(* Logix 5000 project; controller Joltek_RA_5069PLC002 vendor 1 type 14 code 226 rev 34.15; software revision 34.04 *)

TASK MainTask (continuous, watchdog 500 ms) : MainProgram
TASK SafetyTask (periodic, rate 20 ms, priority 10, watchdog 20 ms, safety) : SafetyProgram

MODULES
   Local : vendor 1 type 14 code 226 (5069 0, rev 34.15)
      Joltek_SW001 : vendor 1 type 12 code 231 (Ethernet 192.168.1.70, rev 13.8, Output RPI 1000 ms)
END_MODULES

TYPE UDT_ErrorDataLog :
STRUCT
   Time : UDT_Timestamp;
   DINTlog : DINT[10];
   REALlog : REAL[10];
END_STRUCT
END_TYPE

TYPE UDT_Line :
STRUCT
   Filler : UDT_Machine;
   Capper : UDT_Machine;
   Labeler : UDT_Machine;
   CasePAcker : UDT_Machine;
END_STRUCT
END_TYPE

TYPE UDT_Machine :
STRUCT
   Status : INT;
   Running : TIMER;
   Running_B : BOOL;
   CustomData : DINT[10];
   CustomREALData : REAL[10];
   Faulted : DINT;
END_STRUCT
END_TYPE

TYPE UDT_Timestamp :
STRUCT
   Year : DINT;
   Month : DINT;
   Day : DINT;
   Hour : DINT;
   Minute : DINT;
   Second : DINT;
END_STRUCT
END_TYPE

VAR_GLOBAL   (* controller tags *)
   FillerData : UDT_Machine;
   HMI_BOOL1 : BOOL[128] := ([0] := 1);
        [2]   // Filler - HMI | Station 1 Filling
        [3]   // Filler - HMI | Station 2 Filling
   HMI_INT : INT[100] := ([0] := 3, [1] := 717, [2] := 50, [3] := 16656, [5] := 10, [10] := 3, [11] := 85, [12] := 164, [14] := 9, [20] := 4, [21] := 115, [22] := 5, [23] := 9, [30] := 2, [31] := 66, [33] := 4100, [40] := 2, [41] := 8, [42] := 38, [50] := 4);
        [3].12   // Filler - Start Permissive
        [3].13   // Filler HMI - Start Command
        [23].0   // Labeler - Labeling in Process
        [23].1   // Labeler - Start Permissive
        [23].2   // Labeler - HMI Start Command
        [23].3   // Labeler - Stop Permissive
        [23].4   // Labeler - HMI Stop Command
        [23].5   // Labeler - HMI Faulted Status
        [23].6   // Labeler - HMI Fault Reset Command
        [33].0   // Case Packer - HMI | Case Folding in Progress
        [33].1   // Case Packer - HMI | Case Gluing in Progress
        [33].10   // Case Packer - HMI | Start Permissive
        [33].11   // Case Packer - HMI | Start Command
        [33].12   // Case Packer - HMI | Stop Permissive
        [33].13   // Case Packer - HMI | Stop Command
        [33].15   // Case Packer - HMI | Clear Fault Command
        [41].0   // Palletizer - HMI | Currently Palletizing
        [41].1   // Palletizer - HMI | Start Permissive
        [41].2   // Palletizer - HMI | Start Command
        [41].7   // Palletizer - HMI | Clear Pallet Command
        [50].0   // Line - HIM | Start Permissive
        [50].1   // Line - HIM | Start Command
        [50].2   // Line - HIM | Stop Permissive
        [50].3   // Line - HIM | Stop Command
        [50].5   // Line - HIM | Fault Reset Command
        [14].2   // Capper - HMI | Start Command
        [14].4   // Capper - HMI | Stop Command
        [14].6   // Capper - HMI | Fault Reset Command
   HMI_REAL : REAL[100] := ([0] := 100.0, [1] := 100.0, [2] := 100.0, [3] := 60.0, [4] := 42.0);
   Line1 : UDT_Line;
   Line34Pump3Motor342DischargeOfTank23_Sig : DINT;
   Line45Pump3MTR345InfeedRawIngredientFlou : DINT;
   Line6Pump1DischargeOfTank3 : DINT;
   Sys_DINT : DINT[100] := ([0] := 3, [1] := 3387, [2] := 6708, [3] := 68, [4] := 717, [5] := 10000, [6] := 10000, [7] := 1, [8] := 1, [9] := 1, [10] := 1, [11] := 1, [12] := 1, [13] := 1, [14] := 1, [15] := 1, [16] := 1, [17] := 1, [18] := 1, [19] := 1, [20] := 1, [21] := 1, [22] := 1, [23] := 1, [24] := 1, [25] := 1, [26] := 1, [27] := 1, [28] := 1, [29] := 1, [30] := 1, [31] := 1, [32] := 1, [33] := 1, [34] := 1, [35] := 1, [36] := 1, [39] := 50, [40] := 52, [41] := 10000, [42] := 85, [43] := 164, [44] := 20, [45] := 6100, [46] := 5, [47] := 115, [48] := 4, [49] := 66, [51] := 4200, [54] := 1, [55] := 4, [57] := 38);
        [0]   // Line 1 Motor 324 of the Conveyor 23 Discharge Pump 4-20mA Signal
        [1]   // Line 2 Motor 32334 of the Conveyor 2233 Discharge Pump 0-20mA Signal SCALED
        [3].1   // Filler - Stop
        [3].3   // Filler - Faulted
        [3].2   // Filler - Running
        [40].4   // Capper - Start Capping Process
        [4]   // Filler - Infeed Empty Bottle Count
        [3].0   // Filler - Start
        [3].4   // Filler - Alarm | Infeed Empty Bottle Conveyor Empty
        [3].5   // Filler - Alarm | Infeed Empty Bottle Conveyor Low
        [3].6   // Filler - Alarm | Discharge Filled Bottle Conveyor Full
        [3].7   // Filler - Alarm | Discharge Filled Bottle Conveyor Almost Full
        [40].2   // Capper - Running
        [40].5   // Capper Discharge Conveyor Full
        [40].6   // Capper Discharge Conveyor Almost Full
        [40].7   // Capper Infeed Conveyor Empty
        [40].8   // Capper Infeed Conveyor Almost Empty
        [44].0   // Labeler - Start
        [44].2   // Labeler - Running
        [39]   // Filled Bottle Conveyor Count
        [44].1   // Labeler - Stop
        [44].3   // Labeler - Faulted
        [43]   // Capper - Caps available in the hopper
        [44].5   // Labeler - Labeled Bottle Conveyor Full
        [44].6   // Labeler - Labeled Bottle Conveyor Almost Full
        [44].7   // Labeler - Capped Bottle Conveyor Empty
        [44].8   // Labeler - Capped Bottle Conveyor Almost Empty
        [44].9   // Labeler - Unwind Station Empty
        [44].10   // Labeler - Unwind Station Almost Empty
        [48].0   // Case Packer - Start
        [48].1   // Case Packer - Stop
        [48].3   // Case Packer - Faulted
        [48].2   // Case Packer - Running
        [48].4   // Case Packer - Case Filling Station
        [46]   // Labeled Bollte Conveyor Count
        [49]   // Case Packer - Empty Case Count
        [48].5   // Case Packer - Gluing Station Case in Place
        [48].6   // Case Packer - Case Filled Ready
        [51]   // Case Packer - Glue Station Level (10,000)
        [48].7   // Case Packer - Gluing Station Case Start
        [54].0   // Case Packer - Infeed Labeled Bottles Empty
        [54].1   // Case Packer - Infeed Labeled Bottles Low
        [54].2   // Case Packer - Cases Empty
        [54].3   // Case Packer - Cases Low
        [54].4   // Case Packer - Glue Tank Empty
        [54].5   // Case Packer - Glue Tank Low
        [54].6   // Case Packer - Discharge Conveyor Full
        [54].7   // Case Packer - Discharge Conveyor Almost Full
        [55].0   // Palletizer - Start
        [55].1   // Palletizer - Stop
        [55].3   // Palletizer - Faulted
        [55].2   // Palletizer - Running
        [55].4   // Palletizer - Case Placed by Robot
        [40].0   // Capper - Start
        [40].1   // Capper - Stop
        [40].3   // Capper - Faulted
   Sys_FIFO_C : CONTROL[10] := ([0].LEN := 32, [0].POS := 32, [0].DN := 1);
   Sys_Timer : TIMER[100] := ([0].PRE := 50, [0].ACC := 28, [0].EN := 1, [0].TT := 1, [1].PRE := 150, [1].ACC := 28, [1].EN := 1, [1].TT := 1, [2].PRE := 2000, [2].ACC := 2000, [2].EN := 1, [2].DN := 1, [3].PRE := 200, [3].ACC := 135, [3].EN := 1, [3].TT := 1, [4].PRE := 200, [4].ACC := 135, [4].EN := 1, [4].TT := 1, [10].PRE := 200, [10].ACC := 84, [10].EN := 1, [10].TT := 1, [11].PRE := 50, [11].ACC := 34, [11].EN := 1, [11].TT := 1, [12].PRE := 50, [13].PRE := 100, [14].PRE := 50);
   System_Date_Time : DINT[7] := ([0] := 2026, [1] := 1, [2] := 6, [4] := 14, [5] := 43, [6] := 306763);
   Test_Bool : BOOL[64];
   TestBOOL : BOOL;
   TestControl : CONTROL;
   TestCounter : COUNTER;
   TestDINT : DINT;
   TestDINTArray : DINT[10];
   TestINT : INT;
   TestTimer : TIMER;
   TestTimerArr : TIMER[10];
END_VAR

PROGRAM MainProgram   (* main routine MainRoutine *)
VAR
   CurrentPos1 : DINT := 12;
   Vlad_Test : BOOL[64] := ([0] := 1);
END_VAR

ROUTINE _01_System   (* ladder *)
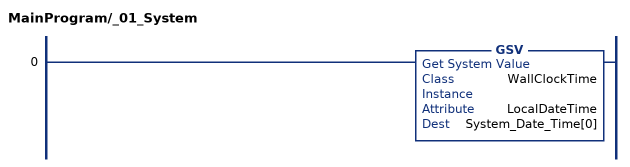
   0: GSV(WallClockTime,,LocalDateTime,System_Date_Time[0]);
END_ROUTINE

ROUTINE _02_Filler   (* ladder *)
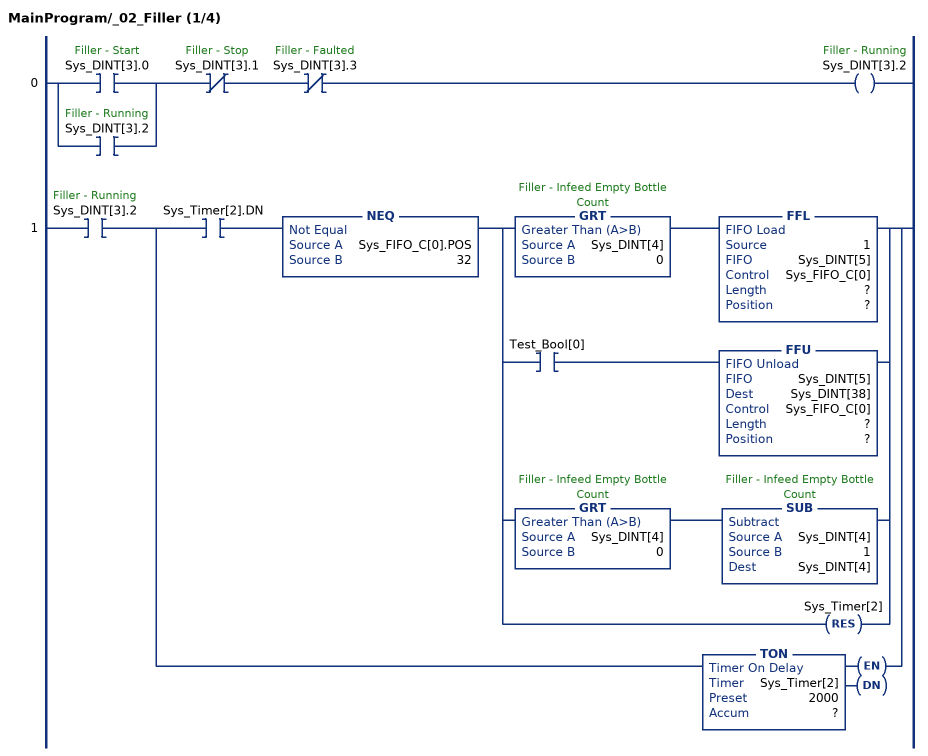
   0: [XIC(Sys_DINT[3].0) ,XIC(Sys_DINT[3].2) ]XIO(Sys_DINT[3].1)XIO(Sys_DINT[3].3)OTE(Sys_DINT[3].2);
   1: XIC(Sys_DINT[3].2)[XIC(Sys_Timer[2].DN) NEQ(Sys_FIFO_C[0].POS,32) [GRT(Sys_DINT[4],0) FFL(1,Sys_DINT[5],Sys_FIFO_C[0],?,?) ,XIC(Test_Bool[0]) FFU(Sys_DINT[5],Sys_DINT[38],Sys_FIFO_C[0],?,?) ,GRT(Sys_DINT[4],0) SUB(Sys_DINT[4],1,Sys_DINT[4]) ,RES(Sys_Timer[2]) ] ,TON(Sys_Timer[2],?,?) ];
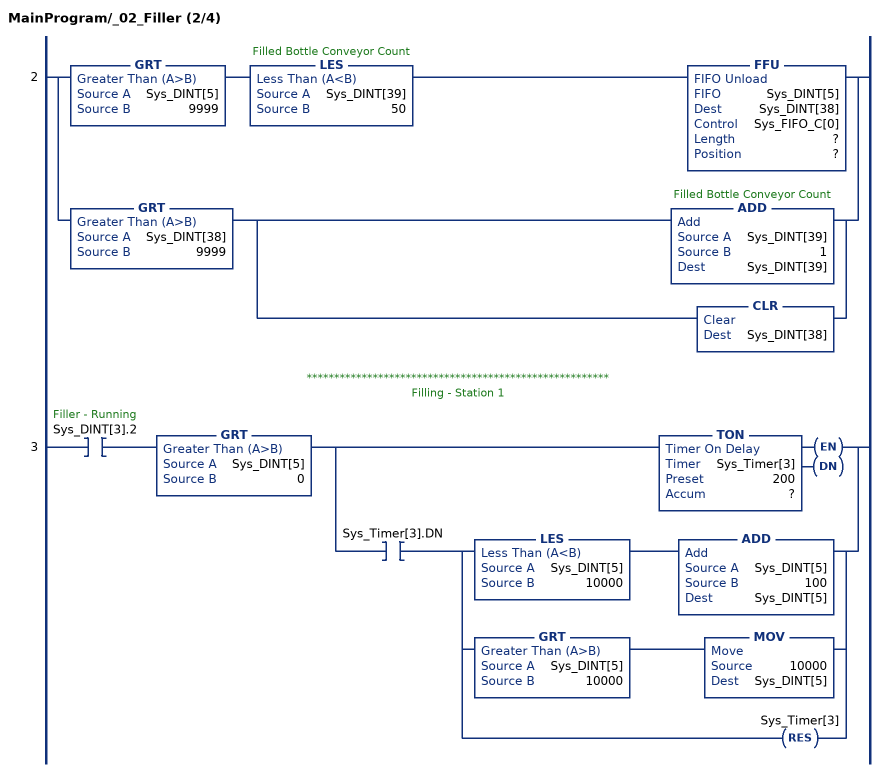
   2: [GRT(Sys_DINT[5],9999) LES(Sys_DINT[39],50) FFU(Sys_DINT[5],Sys_DINT[38],Sys_FIFO_C[0],?,?) ,GRT(Sys_DINT[38],9999) [ADD(Sys_DINT[39],1,Sys_DINT[39]) ,CLR(Sys_DINT[38]) ] ];
   // *******************************************************
   // Filling - Station 1
   3: XIC(Sys_DINT[3].2)GRT(Sys_DINT[5],0)[TON(Sys_Timer[3],?,?) ,XIC(Sys_Timer[3].DN) [LES(Sys_DINT[5],10000) ADD(Sys_DINT[5],100,Sys_DINT[5]) ,GRT(Sys_DINT[5],10000) MOV(10000,Sys_DINT[5]) ,RES(Sys_Timer[3]) ] ];
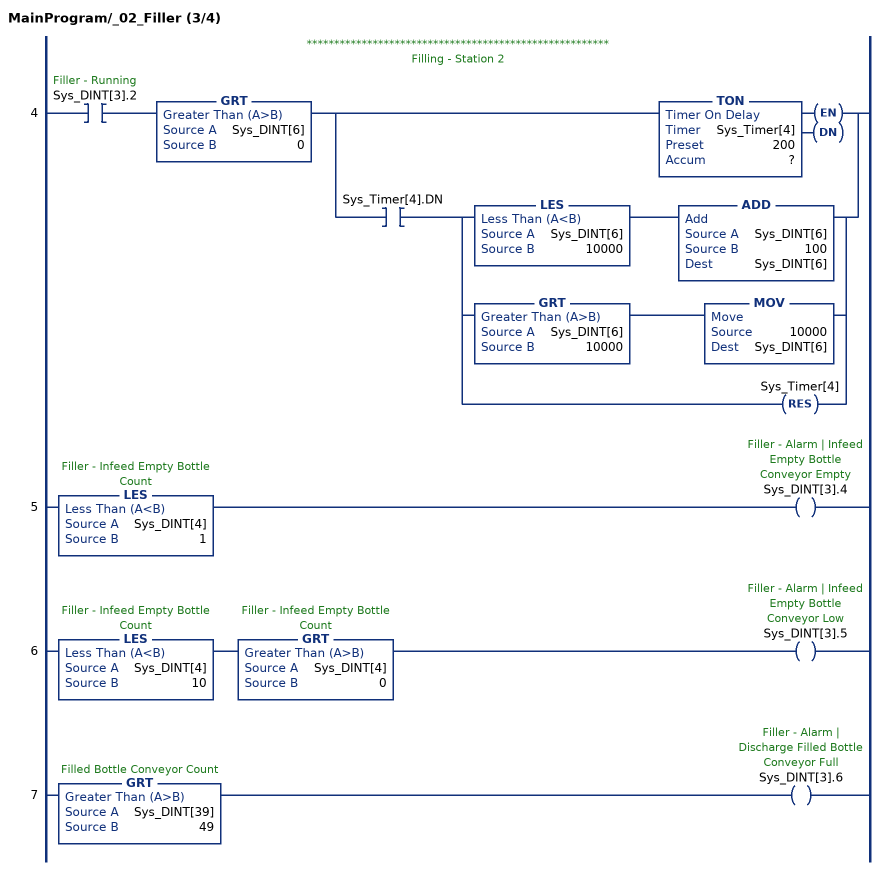
   // *******************************************************
   // Filling - Station 2
   4: XIC(Sys_DINT[3].2)GRT(Sys_DINT[6],0)[TON(Sys_Timer[4],?,?) ,XIC(Sys_Timer[4].DN) [LES(Sys_DINT[6],10000) ADD(Sys_DINT[6],100,Sys_DINT[6]) ,GRT(Sys_DINT[6],10000) MOV(10000,Sys_DINT[6]) ,RES(Sys_Timer[4]) ] ];
   5: LES(Sys_DINT[4],1)OTE(Sys_DINT[3].4);
   6: LES(Sys_DINT[4],10)GRT(Sys_DINT[4],0)OTE(Sys_DINT[3].5);
   7: GRT(Sys_DINT[39],49)OTE(Sys_DINT[3].6);
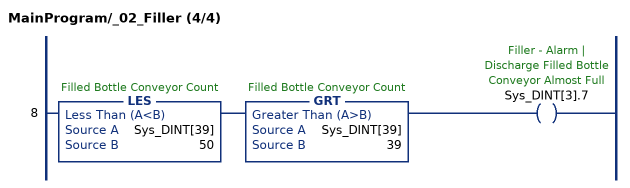
   8: LES(Sys_DINT[39],50)GRT(Sys_DINT[39],39)OTE(Sys_DINT[3].7);
END_ROUTINE

ROUTINE _03_Capper   (* ladder *)
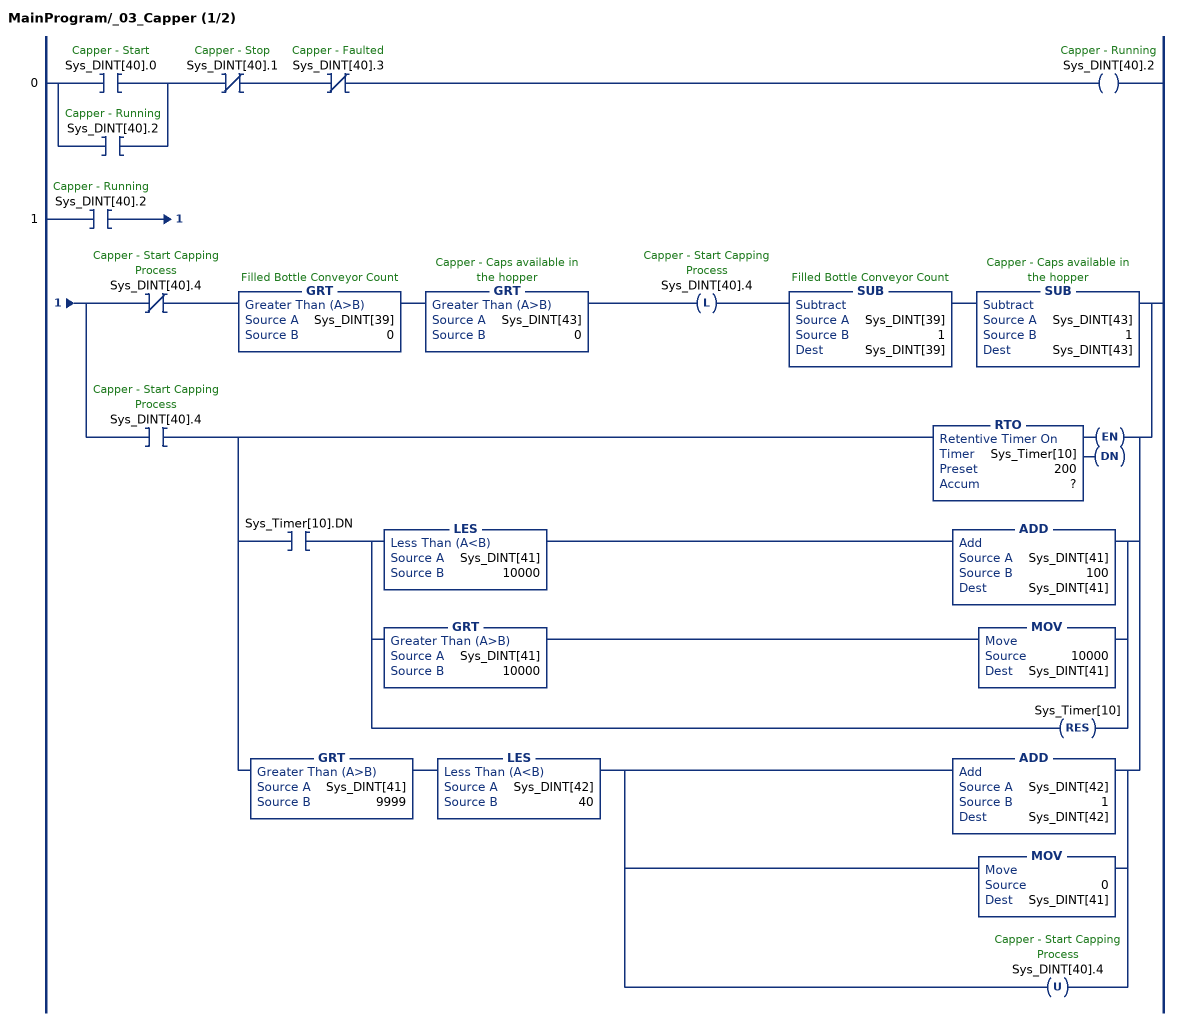
   0: [XIC(Sys_DINT[40].0) ,XIC(Sys_DINT[40].2) ]XIO(Sys_DINT[40].1)XIO(Sys_DINT[40].3)OTE(Sys_DINT[40].2);
   1: XIC(Sys_DINT[40].2)[XIO(Sys_DINT[40].4) GRT(Sys_DINT[39],0) GRT(Sys_DINT[43],0) OTL(Sys_DINT[40].4) SUB(Sys_DINT[39],1,Sys_DINT[39]) SUB(Sys_DINT[43],1,Sys_DINT[43]) ,XIC(Sys_DINT[40].4) [RTO(Sys_Timer[10],?,?) ,XIC(Sys_Timer[10].DN) [LES(Sys_DINT[41],10000) ADD(Sys_DINT[41],100,Sys_DINT[41]) ,GRT(Sys_DINT[41],10000) MOV(10000,Sys_DINT[41]) ,RES(Sys_Timer[10]) ] ,GRT(Sys_DINT[41],9999) LES(Sys_DINT[42],40) [ADD(Sys_DINT[42],1,Sys_DINT[42]) ,MOV(0,Sys_DINT[41]) ,OTU(Sys_DINT[40].4) ] ] ];
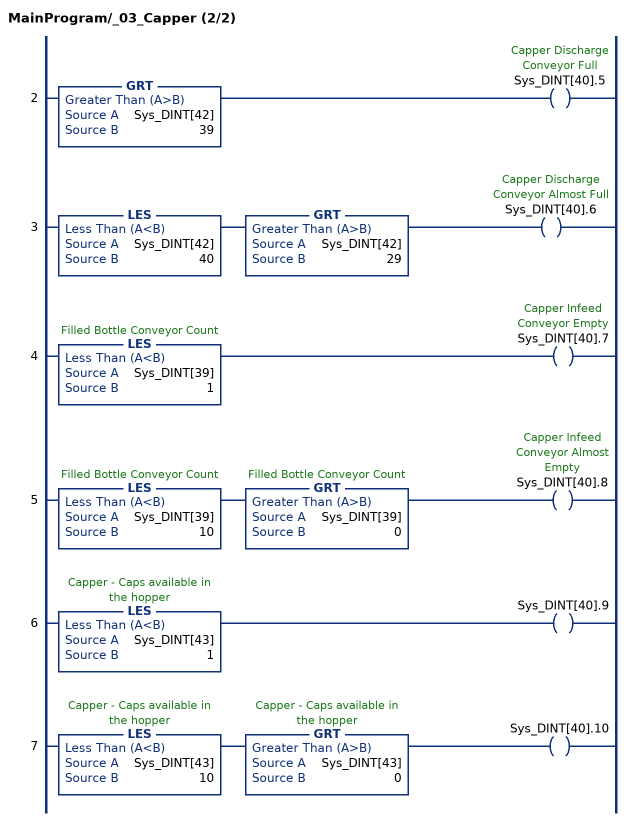
   2: GRT(Sys_DINT[42],39)OTE(Sys_DINT[40].5);
   3: LES(Sys_DINT[42],40)GRT(Sys_DINT[42],29)OTE(Sys_DINT[40].6);
   4: LES(Sys_DINT[39],1)OTE(Sys_DINT[40].7);
   5: LES(Sys_DINT[39],10)GRT(Sys_DINT[39],0)OTE(Sys_DINT[40].8);
   6: LES(Sys_DINT[43],1)OTE(Sys_DINT[40].9);
   7: LES(Sys_DINT[43],10)GRT(Sys_DINT[43],0)OTE(Sys_DINT[40].10);
END_ROUTINE

ROUTINE _04_Labeler   (* ladder *)
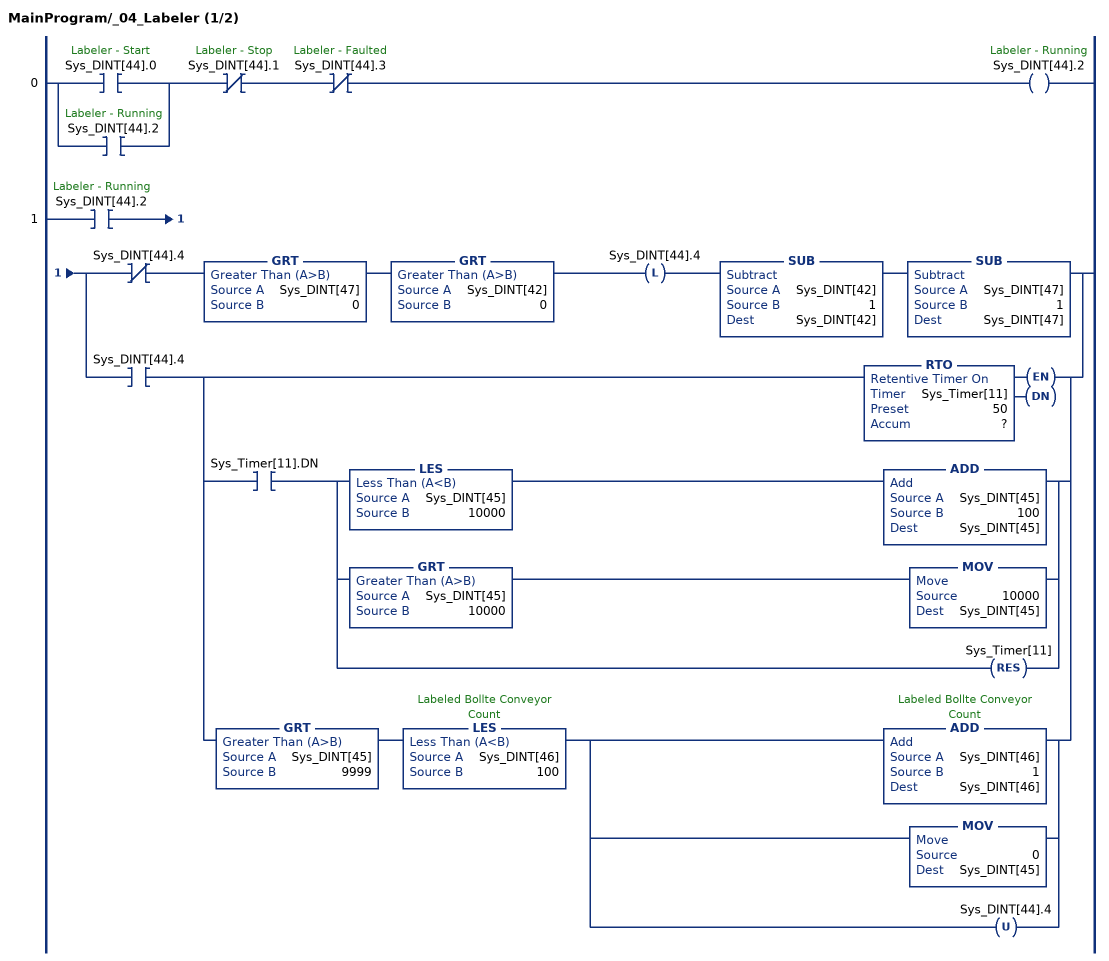
   0: [XIC(Sys_DINT[44].0) ,XIC(Sys_DINT[44].2) ]XIO(Sys_DINT[44].1)XIO(Sys_DINT[44].3)OTE(Sys_DINT[44].2);
   1: XIC(Sys_DINT[44].2)[XIO(Sys_DINT[44].4) GRT(Sys_DINT[47],0) GRT(Sys_DINT[42],0) OTL(Sys_DINT[44].4) SUB(Sys_DINT[42],1,Sys_DINT[42]) SUB(Sys_DINT[47],1,Sys_DINT[47]) ,XIC(Sys_DINT[44].4) [RTO(Sys_Timer[11],?,?) ,XIC(Sys_Timer[11].DN) [LES(Sys_DINT[45],10000) ADD(Sys_DINT[45],100,Sys_DINT[45]) ,GRT(Sys_DINT[45],10000) MOV(10000,Sys_DINT[45]) ,RES(Sys_Timer[11]) ] ,GRT(Sys_DINT[45],9999) LES(Sys_DINT[46],100) [ADD(Sys_DINT[46],1,Sys_DINT[46]) ,MOV(0,Sys_DINT[45]) ,OTU(Sys_DINT[44].4) ] ] ];
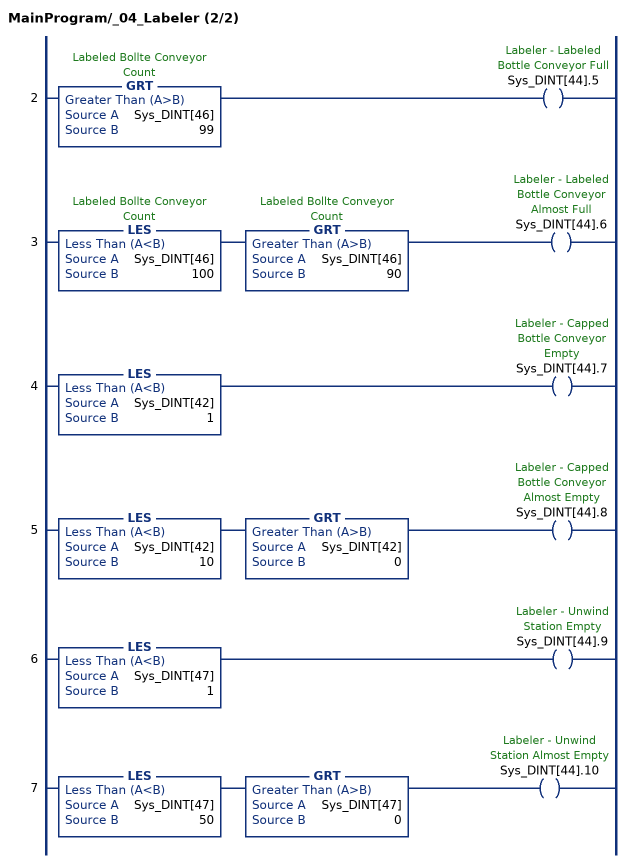
   2: GRT(Sys_DINT[46],99)OTE(Sys_DINT[44].5);
   3: LES(Sys_DINT[46],100)GRT(Sys_DINT[46],90)OTE(Sys_DINT[44].6);
   4: LES(Sys_DINT[42],1)OTE(Sys_DINT[44].7);
   5: LES(Sys_DINT[42],10)GRT(Sys_DINT[42],0)OTE(Sys_DINT[44].8);
   6: LES(Sys_DINT[47],1)OTE(Sys_DINT[44].9);
   7: LES(Sys_DINT[47],50)GRT(Sys_DINT[47],0)OTE(Sys_DINT[44].10);
END_ROUTINE

ROUTINE _05_CasePacker   (* ladder *)
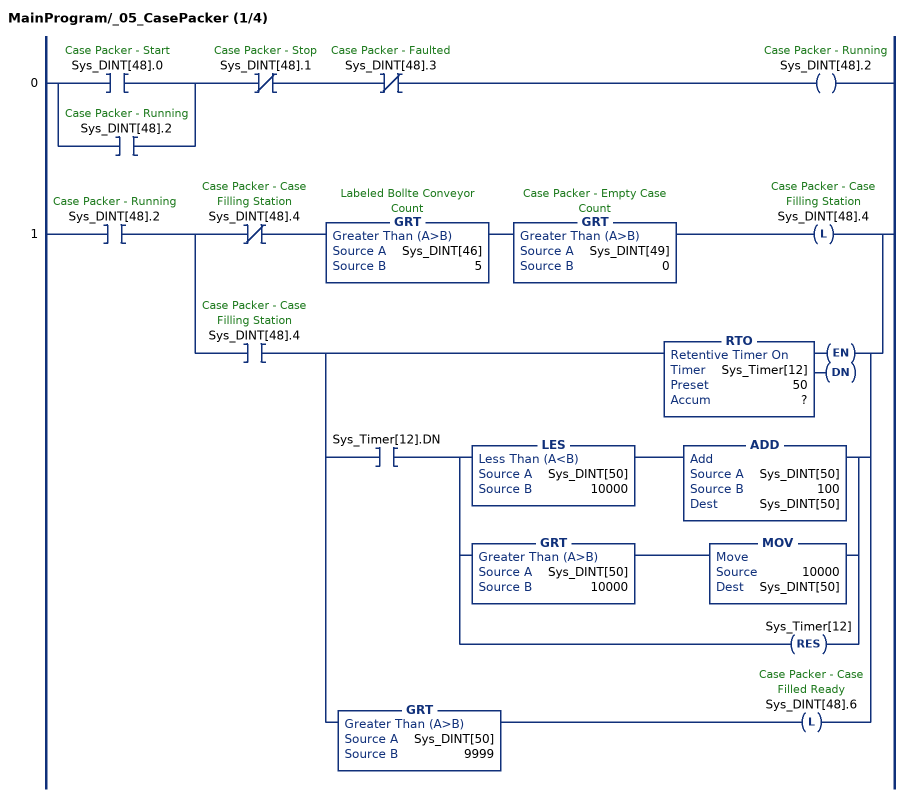
   0: [XIC(Sys_DINT[48].0) ,XIC(Sys_DINT[48].2) ]XIO(Sys_DINT[48].1)XIO(Sys_DINT[48].3)OTE(Sys_DINT[48].2);
   1: XIC(Sys_DINT[48].2)[XIO(Sys_DINT[48].4) GRT(Sys_DINT[46],5) GRT(Sys_DINT[49],0) OTL(Sys_DINT[48].4) ,XIC(Sys_DINT[48].4) [RTO(Sys_Timer[12],?,?) ,XIC(Sys_Timer[12].DN) [LES(Sys_DINT[50],10000) ADD(Sys_DINT[50],100,Sys_DINT[50]) ,GRT(Sys_DINT[50],10000) MOV(10000,Sys_DINT[50]) ,RES(Sys_Timer[12]) ] ,GRT(Sys_DINT[50],9999) OTL(Sys_DINT[48].6) ] ];